// TIA Portal project "ITALTERM_V2.2" (V15)

(* hardware
DEVICE "SIMATIC 1200 station_3"  S71200.Device
   slot 0: "S7-1200 rack"  Rack  V1.0
   slot 1: "MEDIDOR_ITALTERM"  CPU 1214C AC/DC/Rly  6ES7 214-1BG40-0XB0  V4.2
   slot 2: "DI8 x 24VDC / DQ8 x relay_1"  SM 1223 DI16/DQ16 x relay  6ES7 223-1PL32-0XB0  V2.0
   slot 101: "CM 1241 (RS422/485)_1"  6ES7 241-1CH32-0XB0  V2.2
*)

// ===== PLC "MEDIDOR_ITALTERM"  CPU 1214C AC/DC/Rly =====

VAR_GLOBAL   // PLC tag table "Default tag table"
   "System_Byte" AT %MB1 : Byte;
   "FirstScan" AT %M1.0 : Bool;
   "DiagStatusUpdate" AT %M1.1 : Bool;
   "AlwaysTRUE" AT %M1.2 : Bool;
   "AlwaysFALSE" AT %M1.3 : Bool;
   "Clock_Byte" AT %MB270 : Byte;
   "Clock_10Hz" AT %M270.0 : Bool;
   "Clock_5Hz" AT %M270.1 : Bool;
   "Clock_2.5Hz" AT %M270.2 : Bool;
   "Clock_2Hz" AT %M270.3 : Bool;
   "Clock_1.25Hz" AT %M270.4 : Bool;
   "Clock_1Hz" AT %M270.5 : Bool;
   "Clock_0.625Hz" AT %M270.6 : Bool;
   "Clock_0.5Hz" AT %M270.7 : Bool;
END_VAR

DATA_BLOCK "ITALTERM_FB_P2"   // DB81
{ S7_Optimized_Access := 'TRUE' }
VERSION : 0.1
// stored: InstanceOfName ITALTERM_FB
"ITALTERM_FB"
BEGIN
END_DATA_BLOCK

DATA_BLOCK "ITALTERM"   // DB208
{ S7_Optimized_Access := 'FALSE' }
VERSION : 0.1
   VAR
      BUFFER_F1 : Array[0..70] of Char;
      BUFFER_F2 : Array[0..70] of Char;
      BUFFER_F3 : Array[0..70] of Char;
      BUFFER_F4 : Array[0..70] of Char;
      BUFFER_F5 : Array[0..70] of Char;
      BUFFER_F6 : Array[0..70] of Char;
      BUFFER_F7 : Array[0..70] of Char;
      BUFFER_F8 : Array[0..70] of Char;
   END_VAR
BEGIN
END_DATA_BLOCK

FUNCTION_BLOCK "ITALTERM_FB"   // FB5, LAD
{ S7_Optimized_Access := 'TRUE' }
VERSION : 0.1
   VAR_INPUT
      LEITURA_CHARS : Array[0..70] of Char;
   END_VAR
   VAR_OUTPUT
      ID : Int;
      HH : Int;
      MM : Int;
      SS : Int;
      TEMPERATURA : Int;
   END_VAR
   VAR_TEMP
      test_ID : Int;
      AUX_STRING_TEMP : String;
      LEITURA_STRING : String;
      test_TEMP : Int;
      AUX_STRING_SS : String;
      AUX_STRING_MM : String;
      AUX_STRING_HH : String;
      AUX_STRING_ID : String;
      test_HH : Int;
      test_MM : Int;
      test_SS : Int;
   END_VAR
BEGIN

REGION Network 1
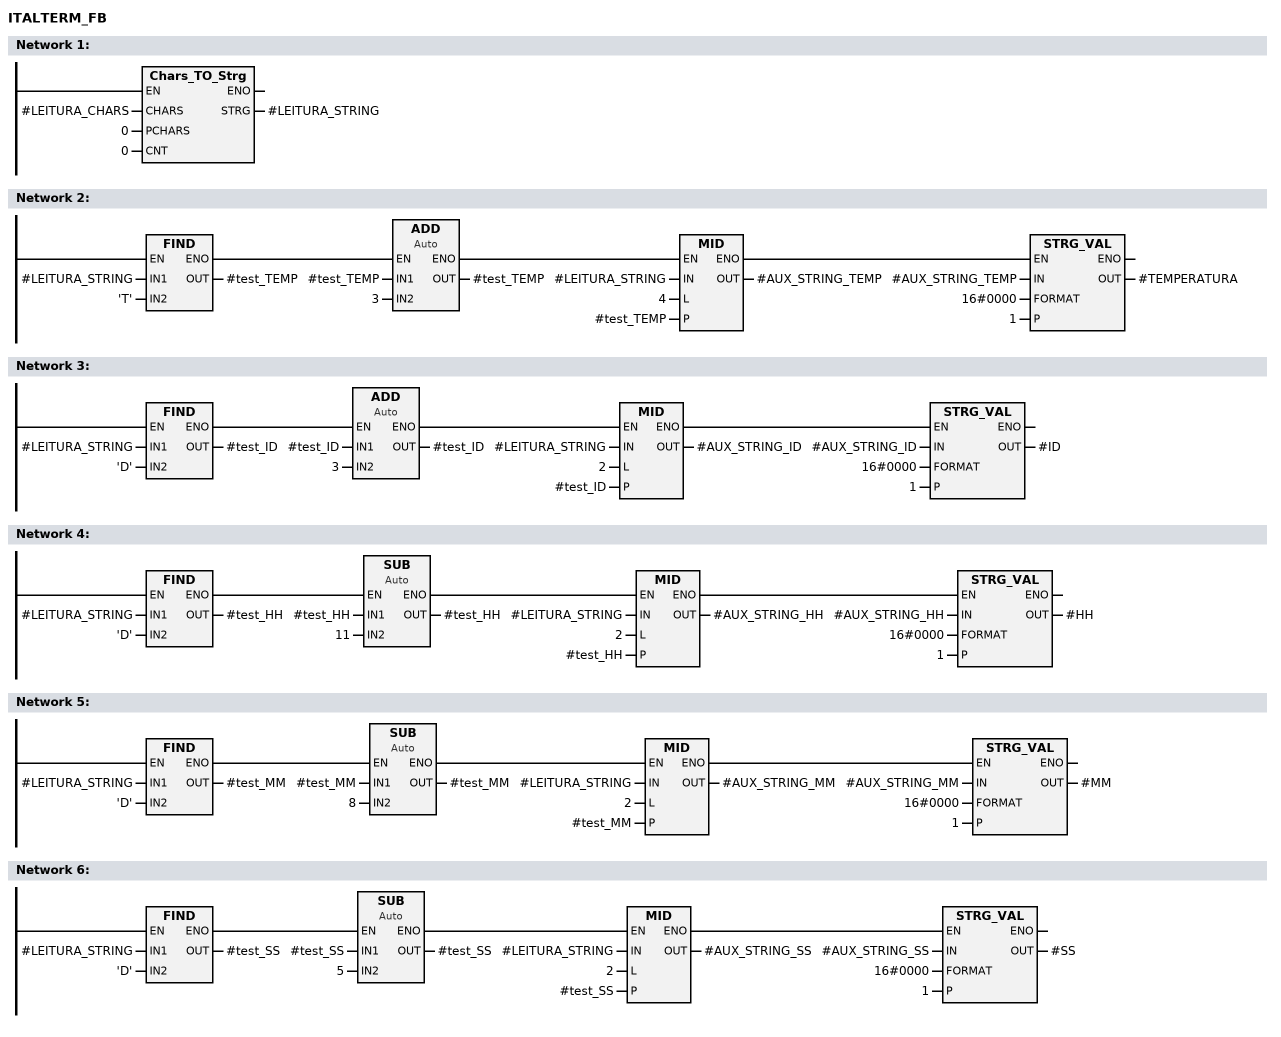
   // no SCL statement known for Chars_TO_Strg: written as a call
   Chars_TO_Strg(Chars := #LEITURA_CHARS, pChars := 0, Cnt := 0, Strg => #LEITURA_STRING);
END_REGION

REGION Network 2
   // ENO of a box is taken as its EN; it also drops when the box reports an error
   #test_TEMP := FIND(IN1 := #LEITURA_STRING, IN2 := 'T');
   #test_TEMP := #test_TEMP + 3;
   #AUX_STRING_TEMP := MID(IN := #LEITURA_STRING, L := 4, P := #test_TEMP);
   STRG_VAL(IN := #AUX_STRING_TEMP, FORMAT := 16#0000, P := 1, OUT => #TEMPERATURA);
END_REGION

REGION Network 3
   // ENO of a box is taken as its EN; it also drops when the box reports an error
   #test_ID := FIND(IN1 := #LEITURA_STRING, IN2 := 'D');
   #test_ID := #test_ID + 3;
   #AUX_STRING_ID := MID(IN := #LEITURA_STRING, L := 2, P := #test_ID);
   STRG_VAL(IN := #AUX_STRING_ID, FORMAT := 16#0000, P := 1, OUT => #ID);
END_REGION

REGION Network 4
   // ENO of a box is taken as its EN; it also drops when the box reports an error
   #test_HH := FIND(IN1 := #LEITURA_STRING, IN2 := 'D');
   #test_HH := #test_HH - 11;
   #AUX_STRING_HH := MID(IN := #LEITURA_STRING, L := 2, P := #test_HH);
   STRG_VAL(IN := #AUX_STRING_HH, FORMAT := 16#0000, P := 1, OUT => #HH);
END_REGION

REGION Network 5
   // ENO of a box is taken as its EN; it also drops when the box reports an error
   #test_MM := FIND(IN1 := #LEITURA_STRING, IN2 := 'D');
   #test_MM := #test_MM - 8;
   #AUX_STRING_MM := MID(IN := #LEITURA_STRING, L := 2, P := #test_MM);
   STRG_VAL(IN := #AUX_STRING_MM, FORMAT := 16#0000, P := 1, OUT => #MM);
END_REGION

REGION Network 6
   // ENO of a box is taken as its EN; it also drops when the box reports an error
   #test_SS := FIND(IN1 := #LEITURA_STRING, IN2 := 'D');
   #test_SS := #test_SS - 5;
   #AUX_STRING_SS := MID(IN := #LEITURA_STRING, L := 2, P := #test_SS);
   STRG_VAL(IN := #AUX_STRING_SS, FORMAT := 16#0000, P := 1, OUT => #SS);
END_REGION
END_FUNCTION_BLOCK

FUNCTION "MEDICAO_TEMPERATURA" : Void   // FC4, LAD
{ S7_Optimized_Access := 'TRUE' }
VERSION : 0.1
   VAR_TEMP
      DONE : Bool;
      BUSY : Bool;
      ERROR : Bool;
      STATUS : Word;
      ERROR_1 : Bool;
      STATU_16 : Word;
      ID_P2 : Int;
      HH : Int;
      MM : Int;
      SS : Int;
      TEMPERATURA : Int;
      aux_time_temp : DInt;
      ULTIMO_MEDIDO : DInt;
   END_VAR
BEGIN

REGION Network 1
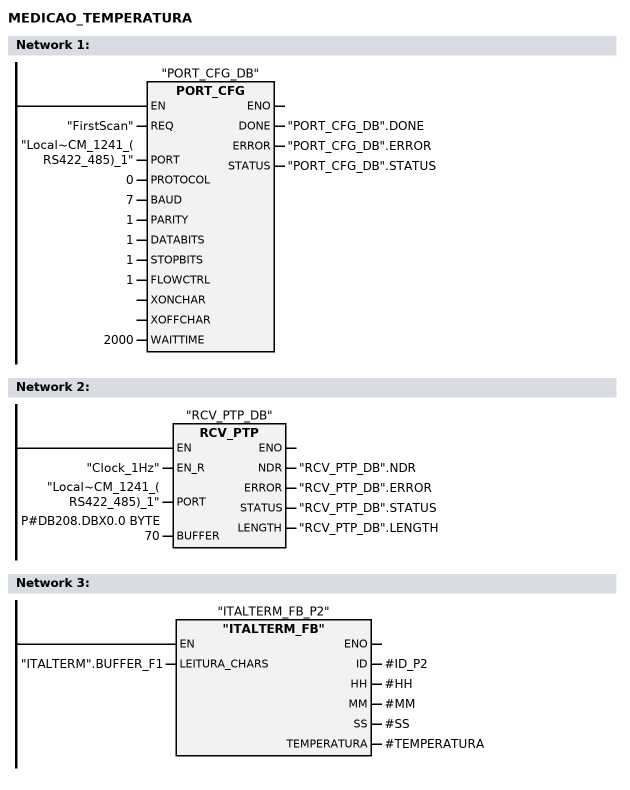
   "PORT_CFG_DB"(REQ := "FirstScan",   // PORT_CFG
                 PORT := "Local~CM_1241_(RS422_485)_1",
                 PROTOCOL := 0,
                 BAUD := 7,
                 PARITY := 1,
                 DATABITS := 1,
                 STOPBITS := 1,
                 FLOWCTRL := 1,
                 WAITTIME := 2000,
                 DONE => "PORT_CFG_DB".DONE,
                 ERROR => "PORT_CFG_DB".ERROR,
                 STATUS => "PORT_CFG_DB".STATUS);
END_REGION

REGION Network 2
   "RCV_PTP_DB"(EN_R := "Clock_1Hz",   // RCV_PTP
                PORT := "Local~CM_1241_(RS422_485)_1",
                BUFFER := P#DB208.DBX0.0 BYTE 70,
                NDR => "RCV_PTP_DB".NDR,
                ERROR => "RCV_PTP_DB".ERROR,
                STATUS => "RCV_PTP_DB".STATUS,
                LENGTH => "RCV_PTP_DB".LENGTH);
END_REGION

REGION Network 3
   RUNG wire#powerrail
      "ITALTERM_FB_P2"(LEITURA_CHARS := "ITALTERM".BUFFER_F1, ID => #ID_P2, HH => #HH, MM => #MM, SS => #SS, TEMPERATURA => #TEMPERATURA)
   END_RUNG
   // the same network as SCL:
   "ITALTERM_FB_P2"(LEITURA_CHARS := "ITALTERM".BUFFER_F1,   // "ITALTERM_FB"
                    ID => #ID_P2,
                    HH => #HH,
                    MM => #MM,
                    SS => #SS,
                    TEMPERATURA => #TEMPERATURA);
END_REGION
END_FUNCTION

ORGANIZATION_BLOCK "Main"   // OB1, LAD, ProgramCycle
TITLE = "Main Program Sweep (Cycle)"
{ S7_Optimized_Access := 'TRUE' }
VERSION : 0.1
   VAR_TEMP
      date_erro : DInt;
      RET : Bool;
      DATA_HORA_ATUAL : DTL;
   END_VAR
BEGIN

REGION Network 1
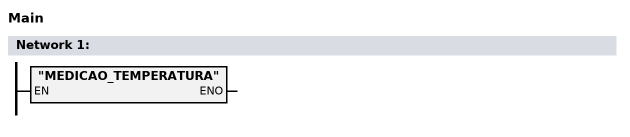
   RUNG wire#powerrail
      "MEDICAO_TEMPERATURA"()
   END_RUNG
   // the same network as SCL:
   "MEDICAO_TEMPERATURA"();
END_REGION
END_ORGANIZATION_BLOCK

(* ===== HMI "HMI_RT_1" =====
connection "HMI_connection_5": 

HMI tags "Default tag table"
   "C" : DInt = PLC SEND."TEMPERATURA MINIMA FORNO 7", 1 s

analog alarms
   11: 'FORNO 6 TEMPERATURA BAIXA', class FORNO 6, trigger "SEND_TEMPERATURA ATUAL FORNO 6"
   12: 'FORNO 6 TEMPERATURA ALTA', class FORNO 6, trigger "SEND_TEMPERATURA ATUAL FORNO 6"
   9: 'FORNO 5 TEMPERATURA BAIXA', class FORNO 5, trigger "SEND_TEMPERATURA ATUAL FORNO 5"
   10: 'FORNO 5 TEMPERATURA ALTA', class FORNO 5, trigger "SEND_TEMPERATURA ATUAL FORNO 5"
   13: 'FORNO 7 TEMPERATURA BAIXA', class FORNO 7, trigger "SEND_TEMPERATURA ATUAL FORNO 7"
   15: 'FORNO 8 TEMPERATURA BAIXA', class FORNO 8, trigger "SEND_TEMPERATURA ATUAL FORNO 8"
   16: 'FORNO 8 TEMPERATURA ALTA', class FORNO 8, trigger "SEND_TEMPERATURA ATUAL FORNO 8"
   14: 'FORNO 7 TEMPERATURA ALTA', class FORNO 7, trigger "SEND_TEMPERATURA ATUAL FORNO 7"
   3: 'FORNO 2 TEMPERATURA BAIXA', class FORNO 2, trigger "SEND_TEMPERATURA ATUAL FORNO 2"
   4: 'FORNO 2 TEMPERATURA ALTA', class FORNO 2, trigger "SEND_TEMPERATURA ATUAL FORNO 2"
   1: 'FORNO 1 TEMPERATURA BAIXA', class FORNO 1, trigger "SEND_TEMPERATURA ATUAL FORNO 1"
   2: 'FORNO 1 TEMPERATURA ALTA', class FORNO 1, trigger "SEND_TEMPERATURA ATUAL FORNO 1"
   7: 'FORNO 4 TEMPERATURA BAIXA', class FORNO 4, trigger "SEND_TEMPERATURA ATUAL FORNO 4"
   8: 'FORNO 4 TEMPERATURA ALTA', class FORNO 4, trigger "SEND_TEMPERATURA ATUAL FORNO 4"
   5: 'FORNO 3 TEMPERATURA BAIXA', class FORNO 3, trigger "SEND_TEMPERATURA ATUAL FORNO 3"
   6: 'FORNO 3 TEMPERATURA ALTA', class FORNO 3, trigger "SEND_TEMPERATURA ATUAL FORNO 3"
   17: 'FORNO 6 TEMPERATURA BAIXA', class FORNO 6, trigger "SEND_TEMPERATURA ATUAL FORNO 6"
   18: 'FORNO 6 TEMPERATURA ALTA', class FORNO 6, trigger "SEND_TEMPERATURA ATUAL FORNO 6"
   19: 'FORNO 5 TEMPERATURA BAIXA', class FORNO 5, trigger "SEND_TEMPERATURA ATUAL FORNO 5"
   20: 'FORNO 5 TEMPERATURA ALTA', class FORNO 5, trigger "SEND_TEMPERATURA ATUAL FORNO 5"
   21: 'FORNO 7 TEMPERATURA BAIXA', class FORNO 7, trigger "SEND_TEMPERATURA ATUAL FORNO 7"
   22: 'FORNO 8 TEMPERATURA BAIXA', class FORNO 8, trigger "SEND_TEMPERATURA ATUAL FORNO 8"
   23: 'FORNO 8 TEMPERATURA ALTA', class FORNO 8, trigger "SEND_TEMPERATURA ATUAL FORNO 8"
   24: 'FORNO 7 TEMPERATURA ALTA', class FORNO 7, trigger "SEND_TEMPERATURA ATUAL FORNO 7"
   25: 'FORNO 2 TEMPERATURA BAIXA', class FORNO 2, trigger "SEND_TEMPERATURA ATUAL FORNO 2"
   26: 'FORNO 2 TEMPERATURA ALTA', class FORNO 2, trigger "SEND_TEMPERATURA ATUAL FORNO 2"
   27: 'FORNO 1 TEMPERATURA BAIXA', class FORNO 1, trigger "SEND_TEMPERATURA ATUAL FORNO 1"
   28: 'FORNO 1 TEMPERATURA ALTA', class FORNO 1, trigger "SEND_TEMPERATURA ATUAL FORNO 1"
   29: 'FORNO 4 TEMPERATURA BAIXA', class FORNO 4, trigger "SEND_TEMPERATURA ATUAL FORNO 4"
   30: 'FORNO 4 TEMPERATURA ALTA', class FORNO 4, trigger "SEND_TEMPERATURA ATUAL FORNO 4"
   31: 'FORNO 3 TEMPERATURA BAIXA', class FORNO 3, trigger "SEND_TEMPERATURA ATUAL FORNO 3"
   32: 'FORNO 3 TEMPERATURA ALTA', class FORNO 3, trigger "SEND_TEMPERATURA ATUAL FORNO 3"

ScreenModuleEditorView "Faceplate_1(1)" 640x480
   StatusForce "Status/Force_1" at 10,10 size 1215x442; ToolTipText 'Text'
*)

(* ===== HMI "HMI_RT_4" =====
system functions are stored by id; their names below are inferred from use

text list "MODO": 0 'DESLIGADO'; 1 'MANUAL'; 2 'AUTOMÁTICO'

text list "MENSAGENS": 0 'SISTEMA OK'

screen "PRINCIPAL_1" 320x240
   TextField "Text field_5" at 67,0 size 186x32; Text 'CONTROLE DOS DUMPERS'
   GraphicView "Graphic view_1" at 253,0 size 67x32; Picture "NOVA LOGO PRI"
   GraphicView "Graphic view" at 0,0 size 67x32; Picture "logos_associadas_logo_whb"
   TextField "Text field_3" at 24,207 size 66x33; Text 'AJUSTE DUMPERS'
   TextField "Text field_2" at 20,45 size 280x30; Text 'MENSAGENS'
   TextField "Text field_4" at 20,125 size 280x30; Text 'MODO OPERAÇÃO'
   SymbolicIOField "Symbolic I/O field_1" at 20,80 size 280x30; TextOff '0'; TextOn '1'; TextList "MENSAGENS"
      ProcessValue <- "DATA_MENSAGENS"
   SymbolicIOField "Symbolic I/O field_2" at 20,160 size 280x30; TextOff '0'; TextOn '1'; TextList "MODO"
      ProcessValue <- "DATA_MODO"
   Softkey "Softkey_F1" at 27,202 size 53x38
      on KeyUp: ActivateScreen("MANUAL DUMPERS AJUSTE", 0)
      on KeyDown: function_b14e0dd5("DATA_MAN-AUTO", 0)
*)